DATA_BLOCK "DB_SDC_EMS_HMI"   // DB3814
{ S7_Optimized_Access := 'FALSE' }
VERSION : 0.1
   VAR
      HEADER : Struct
         DB_NR : Int := 3814;
         Res020 : Int := 0;
         Res040 : Int := 0;
         START_EMS : Int := 20;
         LAENGE_EMS : Int := 260;
         OFFSET_EMS_SEK_STAT : Int := 164;
         LAENGE_EMS_SEK_STAT : Int := 34;
         OFFSET_EMS_FKT : Int := 216;
         START_HMI : Int := 20;
         OFFEST_HMI_DATA : Int := 20;
      END_STRUCT;
      HMI : Array[1..30] of Struct
         PULT_Nr_EDIT : Int;
         BILD_Nr : Int;
         BILD_Nr_Alt : Int;
         EMS_Nr : Int;
         EMS_Nr_Alt : Int;
         PROFIL_Nr : Int;
         PROFIL_Nr_Alt : Int;
         Res140 : Int;
         Res160 : Int;
         T_EDIT : Bool;
         T_RESET_BED : Bool;
         T_SAVE : Bool;
         T_LOAD : Bool;
         Res084 : Bool;
         Res085 : Bool;
         Res086 : Bool;
         Res087 : Bool;
         FR_EDIT : Bool;
         ER_DATA : Bool;
         EMS : "UDT_SDC_EMS";
      END_STRUCT;
   END_VAR
BEGIN
   HMI[1].PULT_Nr_EDIT := 0;
   HMI[1].BILD_Nr := 0;
   HMI[1].BILD_Nr_Alt := 0;
   HMI[1].EMS_Nr := 1;
   HMI[1].EMS_Nr_Alt := 1;
   HMI[1].PROFIL_Nr := 0;
   HMI[1].PROFIL_Nr_Alt := 0;
   HMI[1].Res140 := 0;
   HMI[1].Res160 := 0;
   HMI[1].T_EDIT := FALSE;
   HMI[1].T_RESET_BED := FALSE;
   HMI[1].T_SAVE := FALSE;
   HMI[1].T_LOAD := FALSE;
   HMI[1].Res084 := FALSE;
   HMI[1].Res085 := FALSE;
   HMI[1].Res086 := FALSE;
   HMI[1].Res087 := FALSE;
   HMI[1].FR_EDIT := FALSE;
   HMI[1].ER_DATA := FALSE;
   HMI[1].EMS.IF_I_EMS.STAT.LIFE_BIT := FALSE;
   HMI[1].EMS.IF_I_EMS.STAT.ER_SUM := FALSE;
   HMI[1].EMS.IF_I_EMS.STAT.IR_MAN := TRUE;
   HMI[1].EMS.IF_I_EMS.STAT.ER_RESET := FALSE;
   HMI[1].EMS.IF_I_EMS.STAT.HOIST_CLEAR := FALSE;
   HMI[1].EMS.IF_I_EMS.STAT.POS_START_X := FALSE;
   HMI[1].EMS.IF_I_EMS.STAT.ALWAYS_ONE := TRUE;
   HMI[1].EMS.IF_I_EMS.STAT.H_DISABLED := TRUE;
   HMI[1].EMS.IF_I_EMS.STAT.D_FWD := FALSE;
   HMI[1].EMS.IF_I_EMS.STAT.D_RWD := FALSE;
   HMI[1].EMS.IF_I_EMS.STAT.bit12 := FALSE;
   HMI[1].EMS.IF_I_EMS.STAT.D_IN_POS := TRUE;
   HMI[1].EMS.IF_I_EMS.STAT.H_UP := FALSE;
   HMI[1].EMS.IF_I_EMS.STAT.H_DOWN := FALSE;
   HMI[1].EMS.IF_I_EMS.STAT.H_IN_POS := TRUE;
   HMI[1].EMS.IF_I_EMS.STAT.H_IN_TOPPOS := TRUE;
   HMI[1].EMS.IF_I_EMS.STAT.bit2_0 := FALSE;
   HMI[1].EMS.IF_I_EMS.STAT.bit2_1 := FALSE;
   HMI[1].EMS.IF_I_EMS.STAT.bit2_2 := FALSE;
   HMI[1].EMS.IF_I_EMS.STAT.bit2_3 := TRUE;
   HMI[1].EMS.IF_I_EMS.STAT.IN_BOTPOS := FALSE;
   HMI[1].EMS.IF_I_EMS.STAT.bit2_5 := FALSE;
   HMI[1].EMS.IF_I_EMS.STAT.bit2_6 := FALSE;
   HMI[1].EMS.IF_I_EMS.STAT.bit2_7 := FALSE;
   HMI[1].EMS.IF_I_EMS.STAT.MESS_ACT := TRUE;
   HMI[1].EMS.IF_I_EMS.STAT.MESS_POS := FALSE;
   HMI[1].EMS.IF_I_EMS.STAT.bit3_2 := FALSE;
   HMI[1].EMS.IF_I_EMS.STAT.bit3_3 := FALSE;
   HMI[1].EMS.IF_I_EMS.STAT.bit3_4 := FALSE;
   HMI[1].EMS.IF_I_EMS.STAT.bit3_5 := FALSE;
   HMI[1].EMS.IF_I_EMS.STAT.bit3_6 := FALSE;
   HMI[1].EMS.IF_I_EMS.STAT.DATA_TRANS := TRUE;
   HMI[1].EMS.IF_I_EMS.ERROR := 823;
   HMI[1].EMS.IF_I_EMS.D_POS := 466599;
   HMI[1].EMS.IF_I_EMS.H_POS := 4151;
   HMI[1].EMS.IF_I_EMS.VFC.VFC_No := 16#03;
   HMI[1].EMS.IF_I_EMS.VFC.PW1 := 16#EB40;
   HMI[1].EMS.IF_I_EMS.VFC.PW2 := 16#0000;
   HMI[1].EMS.IF_I_EMS.VFC.PW3 := 16#0000;
   HMI[1].EMS.IF_I_EMS.IQ.BS1PH1_KANAL_1 := FALSE;
   HMI[1].EMS.IF_I_EMS.IQ.BS1PH1_KANAL_2 := FALSE;
   HMI[1].EMS.IF_I_EMS.IQ.BS1PH1_KANAL_3 := FALSE;
   HMI[1].EMS.IF_I_EMS.IQ.BS1PH1_KANAL_4 := FALSE;
   HMI[1].EMS.IF_I_EMS.IQ.BS1PH1_KANAL_5 := FALSE;
   HMI[1].EMS.IF_I_EMS.IQ.BS1PH1_KANAL_6 := FALSE;
   HMI[1].EMS.IF_I_EMS.IQ.BS1PH1_KANAL_7 := FALSE;
   HMI[1].EMS.IF_I_EMS.IQ.BS1PH1_KANAL_8 := FALSE;
   HMI[1].EMS.IF_I_EMS.IQ.BS1FC302 := TRUE;
   HMI[1].EMS.IF_I_EMS.IQ.AB1FCM1 := FALSE;
   HMI[1].EMS.IF_I_EMS.IQ.AB1QA1_R := FALSE;
   HMI[1].EMS.IF_I_EMS.IQ.I_1_3 := FALSE;
   HMI[1].EMS.IF_I_EMS.IQ.I_1_8 := FALSE;
   HMI[1].EMS.IF_I_EMS.IQ.I_1_5 := FALSE;
   HMI[1].EMS.IF_I_EMS.IQ.I_1_6 := FALSE;
   HMI[1].EMS.IF_I_EMS.IQ.I_1_7 := FALSE;
   HMI[1].EMS.IF_I_EMS.IQ.HE1BGS03a := TRUE;
   HMI[1].EMS.IF_I_EMS.IQ.HE1BGS03b := TRUE;
   HMI[1].EMS.IF_I_EMS.IQ.HE1BGS05 := TRUE;
   HMI[1].EMS.IF_I_EMS.IQ.BS1SFWE2 := FALSE;
   HMI[1].EMS.IF_I_EMS.IQ.I_2_4 := FALSE;
   HMI[1].EMS.IF_I_EMS.IQ.I_2_5 := FALSE;
   HMI[1].EMS.IF_I_EMS.IQ.I_2_6 := FALSE;
   HMI[1].EMS.IF_I_EMS.IQ.I_2_7 := FALSE;
   HMI[1].EMS.IF_I_EMS.IQ.I_6_0 := FALSE;
   HMI[1].EMS.IF_I_EMS.IQ.I_6_1 := FALSE;
   HMI[1].EMS.IF_I_EMS.IQ.I_6_2 := FALSE;
   HMI[1].EMS.IF_I_EMS.IQ.I_6_3 := FALSE;
   HMI[1].EMS.IF_I_EMS.IQ.I_6_4 := FALSE;
   HMI[1].EMS.IF_I_EMS.IQ.I_6_5 := FALSE;
   HMI[1].EMS.IF_I_EMS.IQ.I_6_6 := FALSE;
   HMI[1].EMS.IF_I_EMS.IQ.I_6_7 := FALSE;
   HMI[1].EMS.IF_I_EMS.IQ."BS1PH1_L+" := TRUE;
   HMI[1].EMS.IF_I_EMS.IQ.BS1PH1_DAT := FALSE;
   HMI[1].EMS.IF_I_EMS.IQ.AB1QA1 := FALSE;
   HMI[1].EMS.IF_I_EMS.IQ.O_0_3 := FALSE;
   HMI[1].EMS.IF_I_EMS.IQ.O_0_4 := FALSE;
   HMI[1].EMS.IF_I_EMS.IQ.O_0_5 := FALSE;
   HMI[1].EMS.IF_I_EMS.IQ.O_0_6 := FALSE;
   HMI[1].EMS.IF_I_EMS.IQ.O_0_7 := FALSE;
   HMI[1].EMS.IF_I_EMS.IQ.HE1KK1 := FALSE;
   HMI[1].EMS.IF_I_EMS.IQ.O_8_1 := FALSE;
   HMI[1].EMS.IF_I_EMS.IQ.O_8_2 := FALSE;
   HMI[1].EMS.IF_I_EMS.IQ.O_8_3 := FALSE;
   HMI[1].EMS.IF_I_EMS.IQ.O_8_4 := FALSE;
   HMI[1].EMS.IF_I_EMS.IQ.O_8_5 := FALSE;
   HMI[1].EMS.IF_I_EMS.IQ.O_8_6 := FALSE;
   HMI[1].EMS.IF_I_EMS.IQ.O_8_7 := FALSE;
   HMI[1].EMS.IF_I_EMS.IQ.I_261_0 := FALSE;
   HMI[1].EMS.IF_I_EMS.IQ.I_261_1 := FALSE;
   HMI[1].EMS.IF_I_EMS.IQ.I_261_2 := FALSE;
   HMI[1].EMS.IF_I_EMS.IQ.I_261_3 := FALSE;
   HMI[1].EMS.IF_I_EMS.IQ.I_261_4 := FALSE;
   HMI[1].EMS.IF_I_EMS.IQ.I_261_5 := FALSE;
   HMI[1].EMS.IF_I_EMS.IQ.I_261_6 := FALSE;
   HMI[1].EMS.IF_I_EMS.IQ.I_261_7 := FALSE;
   HMI[1].EMS.IF_I_EMS.IQ.HE1BGG1 := TRUE;
   HMI[1].EMS.IF_I_EMS.IQ."HE1BGG1:13" := FALSE;
   HMI[1].EMS.IF_I_EMS.IQ.HE1BGE05 := TRUE;
   HMI[1].EMS.IF_I_EMS.IQ.I_271_3 := FALSE;
   HMI[1].EMS.IF_I_EMS.IQ.I_271_4 := FALSE;
   HMI[1].EMS.IF_I_EMS.IQ.I_271_5 := FALSE;
   HMI[1].EMS.IF_I_EMS.IQ.I_271_6 := FALSE;
   HMI[1].EMS.IF_I_EMS.IQ.I_271_7 := FALSE;
   HMI[1].EMS.IF_I_EMS.IQ.SN1BGE04 := TRUE;
   HMI[1].EMS.IF_I_EMS.IQ.I_281_1 := FALSE;
   HMI[1].EMS.IF_I_EMS.IQ.I_281_2 := FALSE;
   HMI[1].EMS.IF_I_EMS.IQ.I_281_3 := FALSE;
   HMI[1].EMS.IF_I_EMS.IQ.I_281_4 := FALSE;
   HMI[1].EMS.IF_I_EMS.IQ.I_281_5 := FALSE;
   HMI[1].EMS.IF_I_EMS.IQ.I_281_6 := FALSE;
   HMI[1].EMS.IF_I_EMS.IQ.I_281_7 := FALSE;
   HMI[1].EMS.IF_I_EMS.IQ.I_285_0 := FALSE;
   HMI[1].EMS.IF_I_EMS.IQ.I_285_1 := FALSE;
   HMI[1].EMS.IF_I_EMS.IQ.I_285_2 := FALSE;
   HMI[1].EMS.IF_I_EMS.IQ.I_285_3 := FALSE;
   HMI[1].EMS.IF_I_EMS.IQ.I_285_4 := FALSE;
   HMI[1].EMS.IF_I_EMS.IQ.I_285_5 := FALSE;
   HMI[1].EMS.IF_I_EMS.IQ.I_285_6 := FALSE;
   HMI[1].EMS.IF_I_EMS.IQ.I_285_7 := FALSE;
   HMI[1].EMS.IF_I_EMS.ER_WORD_No := 25;
   HMI[1].EMS.IF_I_EMS.ER_WORD := 16#0002;
   HMI[1].EMS.IF_I_EMS.FB_DBNo := 2;
   HMI[1].EMS.IF_I_EMS.FB_DBBNo := 20;
   HMI[1].EMS.IF_Q_EMS.EMS_ID := 1;
   HMI[1].EMS.IF_Q_EMS.CONT.LIFE_BIT := TRUE;
   HMI[1].EMS.IF_Q_EMS.CONT.ER_SDC := FALSE;
   HMI[1].EMS.IF_Q_EMS.CONT.H_EMERG := FALSE;
   HMI[1].EMS.IF_Q_EMS.CONT.Spare_0_3 := FALSE;
   HMI[1].EMS.IF_Q_EMS.CONT.LAMP_TEST := FALSE;
   HMI[1].EMS.IF_Q_EMS.CONT.VAC_CLEAN := FALSE;
   HMI[1].EMS.IF_Q_EMS.CONT.SYNCH := FALSE;
   HMI[1].EMS.IF_Q_EMS.CONT.DATA_TRANS := TRUE;
   HMI[1].EMS.IF_Q_EMS.CONT.ER_RESET := FALSE;
   HMI[1].EMS.IF_Q_EMS.CONT.AUTO := FALSE;
   HMI[1].EMS.IF_Q_EMS.CONT.MAN := TRUE;
   HMI[1].EMS.IF_Q_EMS.CONT.D_C_BREAK := FALSE;
   HMI[1].EMS.IF_Q_EMS.CONT.H_C_BREAK := FALSE;
   HMI[1].EMS.IF_Q_EMS.CONT.D_EMERG_FC := FALSE;
   HMI[1].EMS.IF_Q_EMS.CONT.INC_TOL_POS := FALSE;
   HMI[1].EMS.IF_Q_EMS.CONT.E_STOP := FALSE;
   HMI[1].EMS.IF_Q_EMS.CONT.D_C_FWD := FALSE;
   HMI[1].EMS.IF_Q_EMS.CONT.D_C_RWD := FALSE;
   HMI[1].EMS.IF_Q_EMS.CONT.D_C_BSP := FALSE;
   HMI[1].EMS.IF_Q_EMS.CONT.Spare_2_3 := FALSE;
   HMI[1].EMS.IF_Q_EMS.CONT.IR_noEMSnumber := FALSE;
   HMI[1].EMS.IF_Q_EMS.CONT.IR_noLogin := FALSE;
   HMI[1].EMS.IF_Q_EMS.CONT.BYP_scalance_PN_error := FALSE;
   HMI[1].EMS.IF_Q_EMS.CONT.Spare_2_7 := FALSE;
   HMI[1].EMS.IF_Q_EMS.CONT.H_C_UP := FALSE;
   HMI[1].EMS.IF_Q_EMS.CONT.H_C_DOWN := FALSE;
   HMI[1].EMS.IF_Q_EMS.CONT.H_C_POS := FALSE;
   HMI[1].EMS.IF_Q_EMS.CONT.H_C_TOP := FALSE;
   HMI[1].EMS.IF_Q_EMS.CONT.H_EN := TRUE;
   HMI[1].EMS.IF_Q_EMS.CONT.H_BYP_ROPE := FALSE;
   HMI[1].EMS.IF_Q_EMS.CONT.Spare_3_6 := FALSE;
   HMI[1].EMS.IF_Q_EMS.CONT.H_BYP_REF_INI := FALSE;
   HMI[1].EMS.IF_Q_EMS.D_SETPOS := 466601;
   HMI[1].EMS.IF_Q_EMS.D_SETSPEED := 4000;
   HMI[1].EMS.IF_Q_EMS.H_SETPOS := 4151;
   HMI[1].EMS.IF_Q_EMS.H_SETSPEED := 0;
   HMI[1].EMS.IF_Q_EMS.FB_VFC_No := 16#03;
   HMI[1].EMS.IF_Q_EMS.FB_ER_WORD_No := 25;
   HMI[1].EMS.IF_Q_EMS.DB_No := 2;
   HMI[1].EMS.IF_Q_EMS.DBB_No := 24;
   HMI[1].EMS.IF_Q_EMS.DB_UserData := 16#2710_3B1A;
   HMI[1].EMS.IF_Q_EMS.ERRORS_SPLC._901_ER_SUM := FALSE;
   HMI[1].EMS.IF_Q_EMS.ERRORS_SPLC._902_ER_SUM_SDC := FALSE;
   HMI[1].EMS.IF_Q_EMS.ERRORS_SPLC._903_ER_BC_JUMP := FALSE;
   HMI[1].EMS.IF_Q_EMS.ERRORS_SPLC._904_ER_NO_SEK := FALSE;
   HMI[1].EMS.IF_Q_EMS.ERRORS_SPLC._905_ER_COMMAND := FALSE;
   HMI[1].EMS.IF_Q_EMS.ERRORS_SPLC._906_ER_BC_LIM := FALSE;
   HMI[1].EMS.IF_Q_EMS.ERRORS_SPLC._907_ER_EMS_ID := FALSE;
   HMI[1].EMS.IF_Q_EMS.ERRORS_SPLC._908_ER_SEK_NR := FALSE;
   HMI[1].EMS.IF_Q_EMS.ERRORS_SPLC._909_ER_LIFE := FALSE;
   HMI[1].EMS.IF_Q_EMS.ERRORS_SPLC._910_ER_BUS := FALSE;
   HMI[1].EMS.IF_Q_EMS.ERRORS_SPLC._911 := FALSE;
   HMI[1].EMS.IF_Q_EMS.ERRORS_SPLC._912 := FALSE;
   HMI[1].EMS.IF_Q_EMS.ERRORS_SPLC._913 := FALSE;
   HMI[1].EMS.IF_Q_EMS.ERRORS_SPLC._914 := FALSE;
   HMI[1].EMS.IF_Q_EMS.ERRORS_SPLC._915 := FALSE;
   HMI[1].EMS.IF_Q_EMS.ERRORS_SPLC._916 := FALSE;
   // 9920 more start values not shown
END_DATA_BLOCK

DATA_BLOCK "DB_SDC_TS_IF_HMI"   // DB3816
{ S7_Optimized_Access := 'FALSE' }
AUTHOR : FFM
FAMILY : SDC
NAME : SECT_DEF
VERSION : 1.0
   VAR
      HEADER : Struct
         DB_NR : Int := 3816;
         Res020 : Int := 0;
         Res040 : Int := 0;
         START_DAT : Int := 1;
         LAENGE_SEK_COM : Int := 18;
         LAENGE_SEK_STAT : Int := 34;
         OFFEST_SEK_STAT : Int := 18;
         Res140 : Int := 44;
         START_HMI : Int := 20;
         OFFEST_HMI_DATA : Int := 20;
      END_STRUCT;
      HMI : Array[1..30] of Struct
         PULT_Nr_EDIT : Int;
         BILD_Nr : Int;
         BILD_Nr_Alt : Int;
         SEK_Nr : Int;
         SEK_Nr_Alt : Int;
         Res100 : Int;
         Res120 : Int;
         Res140 : Int;
         Res160 : Int;
         T_EDIT : Bool;
         T_RESET_BED : Bool;
         T_SAVE : Bool;
         T_LOAD : Bool;
         Res084 : Bool;
         Res085 : Bool;
         Res086 : Bool;
         Res087 : Bool;
         FR_EDIT : Bool;
         ER_DATA : Bool;
         COM : "UDT_SDC_EMS_TS_COM";
         STAT : "UDT_SDC_EMS_TS_STAT";
      END_STRUCT;
   END_VAR
BEGIN
   HMI[1].PULT_Nr_EDIT := 0;
   HMI[1].BILD_Nr := 0;
   HMI[1].BILD_Nr_Alt := 0;
   HMI[1].SEK_Nr := 1;
   HMI[1].SEK_Nr_Alt := 255;
   HMI[1].Res100 := 0;
   HMI[1].Res120 := 0;
   HMI[1].Res140 := 0;
   HMI[1].Res160 := 0;
   HMI[1].T_EDIT := FALSE;
   HMI[1].T_RESET_BED := FALSE;
   HMI[1].T_SAVE := FALSE;
   HMI[1].T_LOAD := FALSE;
   HMI[1].Res084 := FALSE;
   HMI[1].Res085 := FALSE;
   HMI[1].Res086 := FALSE;
   HMI[1].Res087 := FALSE;
   HMI[1].FR_EDIT := FALSE;
   HMI[1].ER_DATA := FALSE;
   HMI[1].COM.VAL.PROFIL := 0;
   HMI[1].COM.VAL.D_SETSPEED := 0;
   HMI[1].COM.VAL.D_POS_OFFS := 0;
   HMI[1].COM.BIT.ER_RESET := FALSE;
   HMI[1].COM.BIT.AUTO := FALSE;
   HMI[1].COM.BIT.MAN := FALSE;
   HMI[1].COM.BIT.Spare_0_3 := FALSE;
   HMI[1].COM.BIT.Spare_0_4 := FALSE;
   HMI[1].COM.BIT.E_STOP := TRUE;
   HMI[1].COM.BIT.Spare_0_6 := FALSE;
   HMI[1].COM.BIT.Spare_0_7 := FALSE;
   HMI[1].COM.BIT.D_C_FWD := FALSE;
   HMI[1].COM.BIT.D_C_RWD := FALSE;
   HMI[1].COM.BIT.D_C_BSP := FALSE;
   HMI[1].COM.BIT.D_C_V1 := TRUE;
   HMI[1].COM.BIT.D_C_V2 := FALSE;
   HMI[1].COM.BIT.D_C_V_VAR := FALSE;
   HMI[1].COM.BIT.D_C_BEFOR_POS := FALSE;
   HMI[1].COM.BIT.D_C_AFTER_POS := FALSE;
   HMI[1].COM.BIT.H_C_RAISE := FALSE;
   HMI[1].COM.BIT.H_C_LOWER := FALSE;
   HMI[1].COM.BIT.H_C_POS := FALSE;
   HMI[1].COM.BIT.H_C_POS1 := FALSE;
   HMI[1].COM.BIT.H_C_POS2 := FALSE;
   HMI[1].COM.BIT.H_C_POS3 := FALSE;
   HMI[1].COM.BIT.H_C_POS4 := FALSE;
   HMI[1].COM.BIT.H_C_TOP := FALSE;
   HMI[1].COM.BIT.H_BYP_ROPE := FALSE;
   HMI[1].COM.BIT.Spare_3_1 := FALSE;
   HMI[1].COM.BIT.H_BYP_REF_INI := FALSE;
   HMI[1].COM.BIT.H_C_SLOW := FALSE;
   HMI[1].COM.BIT.D_BYP_DIST_CONTR := FALSE;
   HMI[1].COM.BIT.Spare_3_5 := FALSE;
   HMI[1].COM.BIT.Spare_3_6 := FALSE;
   HMI[1].COM.BIT.SET_PROF := FALSE;
   HMI[1].COM.FKT_SET.EMS_TO_REPAIR_1 := FALSE;
   HMI[1].COM.FKT_SET.EMS_TO_REPAIR_2 := FALSE;
   HMI[1].COM.FKT_SET.EMERG_HOIST := FALSE;
   HMI[1].COM.FKT_SET.Reserve_03 := FALSE;
   HMI[1].COM.FKT_SET.EMERG_DRIVE_FC := FALSE;
   HMI[1].COM.FKT_SET.Reserve_05 := FALSE;
   HMI[1].COM.FKT_SET.LAMP_TEST := FALSE;
   HMI[1].COM.FKT_SET.VAC_CLEAN := FALSE;
   HMI[1].COM.FKT_SET.PE_TEST := FALSE;
   HMI[1].COM.FKT_SET.KOHLE_TEST := FALSE;
   HMI[1].COM.FKT_SET.KOM_TEST := FALSE;
   HMI[1].COM.FKT_SET.Reserve_11 := FALSE;
   HMI[1].COM.FKT_SET.Reserve_12 := FALSE;
   HMI[1].COM.FKT_SET.Reserve_13 := FALSE;
   HMI[1].COM.FKT_SET.Reserve_14 := FALSE;
   HMI[1].COM.FKT_SET.Reserve_15 := FALSE;
   HMI[1].COM.FKT_RESET.EMS_TO_REPAIR_1 := FALSE;
   HMI[1].COM.FKT_RESET.EMS_TO_REPAIR_2 := FALSE;
   HMI[1].COM.FKT_RESET.EMERG_HOIST := FALSE;
   HMI[1].COM.FKT_RESET.Reserve_03 := FALSE;
   HMI[1].COM.FKT_RESET.EMERG_DRIVE_FC := FALSE;
   HMI[1].COM.FKT_RESET.Reserve_05 := FALSE;
   HMI[1].COM.FKT_RESET.LAMP_TEST := FALSE;
   HMI[1].COM.FKT_RESET.VAC_CLEAN := FALSE;
   HMI[1].COM.FKT_RESET.PE_TEST := FALSE;
   HMI[1].COM.FKT_RESET.KOHLE_TEST := FALSE;
   HMI[1].COM.FKT_RESET.KOM_TEST := FALSE;
   HMI[1].COM.FKT_RESET.Reserve_11 := FALSE;
   HMI[1].COM.FKT_RESET.Reserve_12 := FALSE;
   HMI[1].COM.FKT_RESET.Reserve_13 := FALSE;
   HMI[1].COM.FKT_RESET.Reserve_14 := FALSE;
   HMI[1].COM.FKT_RESET.Reserve_15 := FALSE;
   HMI[1].STAT.VAL.EMS_ID := 9;
   HMI[1].STAT.VAL.PROFIL := 1;
   HMI[1].STAT.VAL.DRIVE_POS := 27823;
   HMI[1].STAT.VAL.HOIST_POS := 2747;
   HMI[1].STAT.VAL.ERROR := 824;
   HMI[1].STAT.VAL.DRIVE_POS_PERC := 51;
   HMI[1].STAT.VAL.SEK := 255;
   HMI[1].STAT.BIT.PRESENT := TRUE;
   HMI[1].STAT.BIT.ERROR := FALSE;
   HMI[1].STAT.BIT.MAN_IR := FALSE;
   HMI[1].STAT.BIT.MORE_EMS_PRESENT := FALSE;
   HMI[1].STAT.BIT.ER_COMMAND := FALSE;
   HMI[1].STAT.BIT.W_DIST := FALSE;
   HMI[1].STAT.BIT.Spare_0_6 := FALSE;
   HMI[1].STAT.BIT.MESS_ACT := TRUE;
   HMI[1].STAT.BIT.D_MOVING := FALSE;
   HMI[1].STAT.BIT.D_NOT_MOVING := TRUE;
   HMI[1].STAT.BIT.H_MOVING := FALSE;
   HMI[1].STAT.BIT.H_NOT_MOVING := TRUE;
   HMI[1].STAT.BIT.X_MOVING := FALSE;
   HMI[1].STAT.BIT.X_NOT_MOVING := TRUE;
   HMI[1].STAT.BIT.D_IN_POS := TRUE;
   HMI[1].STAT.BIT.Spare_2_1 := FALSE;
   HMI[1].STAT.BIT.D_BEFOR_POS := FALSE;
   HMI[1].STAT.BIT.D_AFTER_POS := FALSE;
   HMI[1].STAT.BIT.D_GR_AP1 := TRUE;
   HMI[1].STAT.BIT.D_SM_AP1 := FALSE;
   HMI[1].STAT.BIT.D_GR_AP2 := TRUE;
   HMI[1].STAT.BIT.D_SM_AP2 := FALSE;
   HMI[1].STAT.BIT.H_IN_POS := TRUE;
   HMI[1].STAT.BIT.H_IN_TOPPOS := FALSE;
   HMI[1].STAT.BIT.H_IN_POS1 := TRUE;
   HMI[1].STAT.BIT.H_IN_POS2 := TRUE;
   HMI[1].STAT.BIT.H_IN_POS3 := TRUE;
   HMI[1].STAT.BIT.H_IN_POS4 := TRUE;
   HMI[1].STAT.BIT.H_GR_POS := FALSE;
   HMI[1].STAT.BIT.H_SM_POS := FALSE;
   HMI[1].STAT.BIT.H_GR_POS1 := FALSE;
   HMI[1].STAT.BIT.H_SM_POS1 := FALSE;
   HMI[1].STAT.BIT.H_GR_POS2 := FALSE;
   HMI[1].STAT.BIT.H_SM_POS2 := FALSE;
   HMI[1].STAT.BIT.H_GR_POS3 := FALSE;
   HMI[1].STAT.BIT.H_SM_POS3 := FALSE;
   HMI[1].STAT.BIT.H_GR_POS4 := FALSE;
   HMI[1].STAT.BIT.H_SM_POS4 := FALSE;
   HMI[1].STAT.BIT.H_BOTTOM_POS := FALSE;
   HMI[1].STAT.BIT.H_DISABLED := FALSE;
   HMI[1].STAT.BIT.H_CLEAR := FALSE;
   HMI[1].STAT.BIT.D_MOVING_FWD := FALSE;
   HMI[1].STAT.BIT.D_MOVING_RWD := FALSE;
   HMI[1].STAT.BIT.D_RESET_AFTER := FALSE;
   HMI[1].STAT.BIT.D_PULK := FALSE;
   HMI[1].STAT.BIT.D_NO_POS := FALSE;
   HMI[1].STAT.SORTE[1] := 'L';
   HMI[1].STAT.SORTE[2] := 'E';
   HMI[1].STAT.SORTE[3] := 'E';
   HMI[1].STAT.SORTE[4] := 'R';
   HMI[1].STAT.FKT.EMS_TO_REPAIR_1 := FALSE;
   HMI[1].STAT.FKT.EMS_TO_REPAIR_2 := FALSE;
   HMI[1].STAT.FKT.EMERG_HOIST := FALSE;
   HMI[1].STAT.FKT.Reserve_03 := FALSE;
   HMI[1].STAT.FKT.EMERG_DRIVE_FC := FALSE;
   HMI[1].STAT.FKT.Reserve_05 := FALSE;
   HMI[1].STAT.FKT.LAMP_TEST := FALSE;
   HMI[1].STAT.FKT.VAC_CLEAN := FALSE;
   HMI[1].STAT.FKT.PE_TEST := FALSE;
   HMI[1].STAT.FKT.KOHLE_TEST := FALSE;
   HMI[1].STAT.FKT.KOM_TEST := FALSE;
   HMI[1].STAT.FKT.Reserve_11 := FALSE;
   HMI[1].STAT.FKT.Reserve_12 := FALSE;
   HMI[1].STAT.FKT.Reserve_13 := FALSE;
   HMI[1].STAT.FKT.Reserve_14 := FALSE;
   HMI[1].STAT.FKT.Reserve_15 := FALSE;
   HMI[1].STAT.SPARE := 16#0000;
   HMI[2].PULT_Nr_EDIT := 0;
   HMI[2].BILD_Nr := 0;
   HMI[2].BILD_Nr_Alt := 0;
   HMI[2].SEK_Nr := 1;
   HMI[2].SEK_Nr_Alt := 262;
   HMI[2].Res100 := 0;
   HMI[2].Res120 := 0;
   HMI[2].Res140 := 0;
   HMI[2].Res160 := 0;
   HMI[2].T_EDIT := FALSE;
   HMI[2].T_RESET_BED := FALSE;
   HMI[2].T_SAVE := FALSE;
   HMI[2].T_LOAD := FALSE;
   HMI[2].Res084 := FALSE;
   HMI[2].Res085 := FALSE;
   HMI[2].Res086 := FALSE;
   HMI[2].Res087 := FALSE;
   HMI[2].FR_EDIT := FALSE;
   HMI[2].ER_DATA := FALSE;
   HMI[2].COM.VAL.PROFIL := 0;
   HMI[2].COM.VAL.D_SETSPEED := 0;
   HMI[2].COM.VAL.D_POS_OFFS := 0;
   HMI[2].COM.BIT.ER_RESET := FALSE;
   HMI[2].COM.BIT.AUTO := TRUE;
   HMI[2].COM.BIT.MAN := FALSE;
   HMI[2].COM.BIT.Spare_0_3 := FALSE;
   HMI[2].COM.BIT.Spare_0_4 := FALSE;
   HMI[2].COM.BIT.E_STOP := FALSE;
   HMI[2].COM.BIT.Spare_0_6 := FALSE;
   HMI[2].COM.BIT.Spare_0_7 := FALSE;
   HMI[2].COM.BIT.D_C_FWD := TRUE;
   HMI[2].COM.BIT.D_C_RWD := FALSE;
   HMI[2].COM.BIT.D_C_BSP := TRUE;
   HMI[2].COM.BIT.D_C_V1 := TRUE;
   HMI[2].COM.BIT.D_C_V2 := FALSE;
   HMI[2].COM.BIT.D_C_V_VAR := FALSE;
   HMI[2].COM.BIT.D_C_BEFOR_POS := TRUE;
   HMI[2].COM.BIT.D_C_AFTER_POS := TRUE;
   HMI[2].COM.BIT.H_C_RAISE := FALSE;
   HMI[2].COM.BIT.H_C_LOWER := FALSE;
   // 3000 more start values not shown
END_DATA_BLOCK

// folder: 06_IDBs

DATA_BLOCK "IDB504_ZONE_5"   // DB13
{ S7_Optimized_Access := 'FALSE' }
VERSION : 0.1
"FB115_FB_Zone"
BEGIN
END_DATA_BLOCK

DATA_BLOCK "IDB501_ZONE_1"   // DB501
{ S7_Optimized_Access := 'FALSE' }
VERSION : 0.1
"FB115_FB_Zone"
BEGIN
END_DATA_BLOCK

DATA_BLOCK "IDB502_ZONE_2"   // DB502
{ S7_Optimized_Access := 'FALSE' }
VERSION : 0.1
"FB115_FB_Zone"
BEGIN
END_DATA_BLOCK

DATA_BLOCK "IDB503_ZONE_3"   // DB503
{ S7_Optimized_Access := 'FALSE' }
VERSION : 0.1
"FB115_FB_Zone"
BEGIN
END_DATA_BLOCK

DATA_BLOCK "IDB504_ZONE_4"   // DB504
{ S7_Optimized_Access := 'FALSE' }
VERSION : 0.1
"FB115_FB_Zone"
BEGIN
END_DATA_BLOCK

DATA_BLOCK "IDB505_ZONE_5"   // DB505
{ S7_Optimized_Access := 'FALSE' }
VERSION : 0.1
"FB115_FB_Zone"
BEGIN
END_DATA_BLOCK

DATA_BLOCK "IDB506_ZONE_6"   // DB506
{ S7_Optimized_Access := 'FALSE' }
VERSION : 0.1
"FB115_FB_Zone"
BEGIN
END_DATA_BLOCK

DATA_BLOCK "IDB543_ZONE_43"   // DB543
{ S7_Optimized_Access := 'FALSE' }
VERSION : 0.1
"FB115_FB_Zone"
BEGIN
END_DATA_BLOCK

DATA_BLOCK "IDB544_ZONE_44"   // DB544
{ S7_Optimized_Access := 'FALSE' }
VERSION : 0.1
"FB115_FB_Zone"
BEGIN
END_DATA_BLOCK

DATA_BLOCK "IDB547_ZONE_47"   // DB547
{ S7_Optimized_Access := 'FALSE' }
VERSION : 0.1
"FB115_FB_Zone"
BEGIN
END_DATA_BLOCK

DATA_BLOCK "IDB548_ZONE_48"   // DB548
{ S7_Optimized_Access := 'FALSE' }
VERSION : 0.1
"FB115_FB_Zone"
BEGIN
END_DATA_BLOCK

DATA_BLOCK "IDB552_ZONE_52"   // DB552
{ S7_Optimized_Access := 'FALSE' }
VERSION : 0.1
"FB115_FB_Zone"
BEGIN
END_DATA_BLOCK

DATA_BLOCK "IDB558_ZONE_58"   // DB558
{ S7_Optimized_Access := 'FALSE' }
VERSION : 0.1
"FB115_FB_Zone"
BEGIN
END_DATA_BLOCK

DATA_BLOCK "IDB600_ZonePositionArrayTrafficCop_DB"   // DB600
{ S7_Optimized_Access := 'FALSE' }
VERSION : 0.1
"FB116_FB_ZonePositionArrayTrafficCop"
BEGIN
END_DATA_BLOCK

DATA_BLOCK "IDB601_MapSDCOut_Carrier_DB"   // DB601
{ S7_Optimized_Access := 'TRUE' }
VERSION : 0.1
"FB117_MapSDCOut_Carrier"
BEGIN
END_DATA_BLOCK

DATA_BLOCK "IDB602_NextCarrierTCopMotionFB"   // DB602
{ S7_Optimized_Access := 'TRUE' }
VERSION : 0.1
"FB111_NextCarrierTCopMotionFB"
BEGIN
END_DATA_BLOCK

DATA_BLOCK "IDB603_FB_ZonePositionArrayTrafficCop_DB"   // DB603
{ S7_Optimized_Access := 'FALSE' }
VERSION : 0.1
"FB116_FB_ZonePositionArrayTrafficCop"
BEGIN
END_DATA_BLOCK

DATA_BLOCK "IDB604_SpacingCheck"   // DB604
{ S7_Optimized_Access := 'TRUE' }
VERSION : 0.1
"FB120_ZoneSpacingCheck"
BEGIN
END_DATA_BLOCK

DATA_BLOCK "IDB605_CARRIER"   // DB605
{ S7_Optimized_Access := 'TRUE' }
VERSION : 0.1
"FB112_Carrier"
BEGIN
END_DATA_BLOCK

DATA_BLOCK "IDB606_FirstCarrierTCopMotionFB"   // DB606
{ S7_Optimized_Access := 'TRUE' }
VERSION : 0.1
"FB110_FirstCarrierTCopMotionFB"
BEGIN
END_DATA_BLOCK

DATA_BLOCK "IDB607_FirstCarrierTCopMotionFB"   // DB607
{ S7_Optimized_Access := 'TRUE' }
VERSION : 0.1
"FB110_FirstCarrierTCopMotionFB"
BEGIN
END_DATA_BLOCK

DATA_BLOCK "IDB608_NextCarrierTCopMotionFB"   // DB608
{ S7_Optimized_Access := 'TRUE' }
VERSION : 0.1
"FB111_NextCarrierTCopMotionFB"
BEGIN
END_DATA_BLOCK

DATA_BLOCK "IDB609_TCMapSDCOutFB"   // DB609
{ S7_Optimized_Access := 'TRUE' }
VERSION : 0.1
"FB118_TCMapSDCOut"
BEGIN
END_DATA_BLOCK

DATA_BLOCK "IDB610_SpacingCheckFB"   // DB610
{ S7_Optimized_Access := 'TRUE' }
VERSION : 0.1
"FB120_ZoneSpacingCheck"
BEGIN
END_DATA_BLOCK

// folder: System blocks/Program resources

DATA_BLOCK "Reset_Timer"   // DB1
{ S7_Optimized_Access := 'TRUE' }
AUTHOR : Simatic
FAMILY : IEC
NAME : IEC_TMR
VERSION : 1.0
"IEC_TIMER"
BEGIN
END_DATA_BLOCK

DATA_BLOCK "C23_Heartbeat_On_Timer"   // DB2
{ S7_Optimized_Access := 'TRUE' }
AUTHOR : Simatic
FAMILY : IEC
NAME : IEC_TMR
VERSION : 1.0
"IEC_TIMER"
BEGIN
END_DATA_BLOCK

DATA_BLOCK "EMS_Heartbeat_On_Timer"   // DB3
{ S7_Optimized_Access := 'TRUE' }
AUTHOR : Simatic
FAMILY : IEC
NAME : IEC_TMR
VERSION : 1.0
"IEC_TIMER"
BEGIN
END_DATA_BLOCK

DATA_BLOCK "C23_Heartbeat_Off_Timer"   // DB5
{ S7_Optimized_Access := 'TRUE' }
AUTHOR : Simatic
FAMILY : IEC
NAME : IEC_TMR
VERSION : 1.0
"IEC_TIMER"
BEGIN
END_DATA_BLOCK

DATA_BLOCK "C22_Heartbeat_On_Timer"   // DB6
{ S7_Optimized_Access := 'TRUE' }
AUTHOR : Simatic
FAMILY : IEC
NAME : IEC_TMR
VERSION : 1.0
"IEC_TIMER"
BEGIN
END_DATA_BLOCK

DATA_BLOCK "EMS_Heartbeat_Off_Timer"   // DB7
{ S7_Optimized_Access := 'TRUE' }
AUTHOR : Simatic
FAMILY : IEC
NAME : IEC_TMR
VERSION : 1.0
"IEC_TIMER"
BEGIN
END_DATA_BLOCK

DATA_BLOCK "C22_Heartbeat_Off_Timer"   // DB9
{ S7_Optimized_Access := 'TRUE' }
AUTHOR : Simatic
FAMILY : IEC
NAME : IEC_TMR
VERSION : 1.0
"IEC_TIMER"
BEGIN
END_DATA_BLOCK

DATA_BLOCK "C21_Heartbeat_On_Timer"   // DB10
{ S7_Optimized_Access := 'TRUE' }
AUTHOR : Simatic
FAMILY : IEC
NAME : IEC_TMR
VERSION : 1.0
"IEC_TIMER"
BEGIN
END_DATA_BLOCK

DATA_BLOCK "C21_Heartbeat_Off_Timer"   // DB12
{ S7_Optimized_Access := 'TRUE' }
AUTHOR : Simatic
FAMILY : IEC
NAME : IEC_TMR
VERSION : 1.0
"IEC_TIMER"
BEGIN
END_DATA_BLOCK

DATA_BLOCK "C24_Heartbeat_On_Timer"   // DB17
{ S7_Optimized_Access := 'TRUE' }
AUTHOR : Simatic
FAMILY : IEC
NAME : IEC_TMR
VERSION : 1.0
"IEC_TIMER"
BEGIN
END_DATA_BLOCK

DATA_BLOCK "C24_Heartbeat_Off_Timer"   // DB18
{ S7_Optimized_Access := 'TRUE' }
AUTHOR : Simatic
FAMILY : IEC
NAME : IEC_TMR
VERSION : 1.0
"IEC_TIMER"
BEGIN
END_DATA_BLOCK

DATA_BLOCK "C25_Heartbeat_On_Timer"   // DB19
{ S7_Optimized_Access := 'TRUE' }
AUTHOR : Simatic
FAMILY : IEC
NAME : IEC_TMR
VERSION : 1.0
"IEC_TIMER"
BEGIN
END_DATA_BLOCK

DATA_BLOCK "C25_Heartbeat_Off_Timer"   // DB20
{ S7_Optimized_Access := 'TRUE' }
AUTHOR : Simatic
FAMILY : IEC
NAME : IEC_TMR
VERSION : 1.0
"IEC_TIMER"
BEGIN
END_DATA_BLOCK

DATA_BLOCK "C26_Heartbeat_On_Timer"   // DB21
{ S7_Optimized_Access := 'TRUE' }
AUTHOR : Simatic
FAMILY : IEC
NAME : IEC_TMR
VERSION : 1.0
"IEC_TIMER"
BEGIN
END_DATA_BLOCK

DATA_BLOCK "C26_Heartbeat_Off_Timer"   // DB22
{ S7_Optimized_Access := 'TRUE' }
AUTHOR : Simatic
FAMILY : IEC
NAME : IEC_TMR
VERSION : 1.0
"IEC_TIMER"
BEGIN
END_DATA_BLOCK

DATA_BLOCK "C27_Heartbeat_On_Timer"   // DB23
{ S7_Optimized_Access := 'TRUE' }
AUTHOR : Simatic
FAMILY : IEC
NAME : IEC_TMR
VERSION : 1.0
"IEC_TIMER"
BEGIN
END_DATA_BLOCK

DATA_BLOCK "C27_Heartbeat_Off_Timer"   // DB24
{ S7_Optimized_Access := 'TRUE' }
AUTHOR : Simatic
FAMILY : IEC
NAME : IEC_TMR
VERSION : 1.0
"IEC_TIMER"
BEGIN
END_DATA_BLOCK

DATA_BLOCK "C28_Heartbeat_On_Timer"   // DB25
{ S7_Optimized_Access := 'TRUE' }
AUTHOR : Simatic
FAMILY : IEC
NAME : IEC_TMR
VERSION : 1.0
"IEC_TIMER"
BEGIN
END_DATA_BLOCK

DATA_BLOCK "C28_Heartbeat_Off_Timer"   // DB26
{ S7_Optimized_Access := 'TRUE' }
AUTHOR : Simatic
FAMILY : IEC
NAME : IEC_TMR
VERSION : 1.0
"IEC_TIMER"
BEGIN
END_DATA_BLOCK

DATA_BLOCK "C29_Heartbeat_On_Timer"   // DB27
{ S7_Optimized_Access := 'TRUE' }
AUTHOR : Simatic
FAMILY : IEC
NAME : IEC_TMR
VERSION : 1.0
"IEC_TIMER"
BEGIN
END_DATA_BLOCK

DATA_BLOCK "C29_Heartbeat_Off_Timer"   // DB28
{ S7_Optimized_Access := 'TRUE' }
AUTHOR : Simatic
FAMILY : IEC
NAME : IEC_TMR
VERSION : 1.0
"IEC_TIMER"
BEGIN
END_DATA_BLOCK

DATA_BLOCK "C30_Heartbeat_On_Timer"   // DB29
{ S7_Optimized_Access := 'TRUE' }
AUTHOR : Simatic
FAMILY : IEC
NAME : IEC_TMR
VERSION : 1.0
"IEC_TIMER"
BEGIN
END_DATA_BLOCK

DATA_BLOCK "C11_Heartbeat_On_Timer"   // DB30
{ S7_Optimized_Access := 'TRUE' }
AUTHOR : Simatic
FAMILY : IEC
NAME : IEC_TMR
VERSION : 1.0
"IEC_TIMER"
BEGIN
END_DATA_BLOCK

DATA_BLOCK "C11_Heartbeat_Off_Timer"   // DB31
{ S7_Optimized_Access := 'TRUE' }
AUTHOR : Simatic
FAMILY : IEC
NAME : IEC_TMR
VERSION : 1.0
"IEC_TIMER"
BEGIN
END_DATA_BLOCK

DATA_BLOCK "C12_Heartbeat_On_Timer"   // DB32
{ S7_Optimized_Access := 'TRUE' }
AUTHOR : Simatic
FAMILY : IEC
NAME : IEC_TMR
VERSION : 1.0
"IEC_TIMER"
BEGIN
END_DATA_BLOCK

DATA_BLOCK "C12_Heartbeat_Off_Timer"   // DB33
{ S7_Optimized_Access := 'TRUE' }
AUTHOR : Simatic
FAMILY : IEC
NAME : IEC_TMR
VERSION : 1.0
"IEC_TIMER"
BEGIN
END_DATA_BLOCK

DATA_BLOCK "C13_Heartbeat_On_Timer"   // DB34
{ S7_Optimized_Access := 'TRUE' }
AUTHOR : Simatic
FAMILY : IEC
NAME : IEC_TMR
VERSION : 1.0
"IEC_TIMER"
BEGIN
END_DATA_BLOCK

DATA_BLOCK "C13_Heartbeat_Off_Timer"   // DB35
{ S7_Optimized_Access := 'TRUE' }
AUTHOR : Simatic
FAMILY : IEC
NAME : IEC_TMR
VERSION : 1.0
"IEC_TIMER"
BEGIN
END_DATA_BLOCK

DATA_BLOCK "C14_Heartbeat_On_Timer"   // DB36
{ S7_Optimized_Access := 'TRUE' }
AUTHOR : Simatic
FAMILY : IEC
NAME : IEC_TMR
VERSION : 1.0
"IEC_TIMER"
BEGIN
END_DATA_BLOCK

DATA_BLOCK "C14_Heartbeat_Off_Timer"   // DB37
{ S7_Optimized_Access := 'TRUE' }
AUTHOR : Simatic
FAMILY : IEC
NAME : IEC_TMR
VERSION : 1.0
"IEC_TIMER"
BEGIN
END_DATA_BLOCK

DATA_BLOCK "C15_Heartbeat_On_Timer"   // DB38
{ S7_Optimized_Access := 'TRUE' }
AUTHOR : Simatic
FAMILY : IEC
NAME : IEC_TMR
VERSION : 1.0
"IEC_TIMER"
BEGIN
END_DATA_BLOCK

DATA_BLOCK "C15_Heartbeat_Off_Timer"   // DB39
{ S7_Optimized_Access := 'TRUE' }
AUTHOR : Simatic
FAMILY : IEC
NAME : IEC_TMR
VERSION : 1.0
"IEC_TIMER"
BEGIN
END_DATA_BLOCK

DATA_BLOCK "C16_Heartbeat_On_Timer"   // DB40
{ S7_Optimized_Access := 'TRUE' }
AUTHOR : Simatic
FAMILY : IEC
NAME : IEC_TMR
VERSION : 1.0
"IEC_TIMER"
BEGIN
END_DATA_BLOCK

DATA_BLOCK "C16_Heartbeat_Off_Timer"   // DB41
{ S7_Optimized_Access := 'TRUE' }
AUTHOR : Simatic
FAMILY : IEC
NAME : IEC_TMR
VERSION : 1.0
"IEC_TIMER"
BEGIN
END_DATA_BLOCK

DATA_BLOCK "C17_Heartbeat_On_Timer"   // DB42
{ S7_Optimized_Access := 'TRUE' }
AUTHOR : Simatic
FAMILY : IEC
NAME : IEC_TMR
VERSION : 1.0
"IEC_TIMER"
BEGIN
END_DATA_BLOCK

DATA_BLOCK "C17_Heartbeat_Off_Timer"   // DB43
{ S7_Optimized_Access := 'TRUE' }
AUTHOR : Simatic
FAMILY : IEC
NAME : IEC_TMR
VERSION : 1.0
"IEC_TIMER"
BEGIN
END_DATA_BLOCK

DATA_BLOCK "C18_Heartbeat_On_Timer"   // DB44
{ S7_Optimized_Access := 'TRUE' }
AUTHOR : Simatic
FAMILY : IEC
NAME : IEC_TMR
VERSION : 1.0
"IEC_TIMER"
BEGIN
END_DATA_BLOCK

DATA_BLOCK "C18_Heartbeat_Off_Timer"   // DB45
{ S7_Optimized_Access := 'TRUE' }
AUTHOR : Simatic
FAMILY : IEC
NAME : IEC_TMR
VERSION : 1.0
"IEC_TIMER"
BEGIN
END_DATA_BLOCK

DATA_BLOCK "C19_Heartbeat_On_Timer"   // DB46
{ S7_Optimized_Access := 'TRUE' }
AUTHOR : Simatic
FAMILY : IEC
NAME : IEC_TMR
VERSION : 1.0
"IEC_TIMER"
BEGIN
END_DATA_BLOCK

DATA_BLOCK "C19_Heartbeat_Off_Timer"   // DB47
{ S7_Optimized_Access := 'TRUE' }
AUTHOR : Simatic
FAMILY : IEC
NAME : IEC_TMR
VERSION : 1.0
"IEC_TIMER"
BEGIN
END_DATA_BLOCK

DATA_BLOCK "C20_Heartbeat_On_Timer"   // DB48
{ S7_Optimized_Access := 'TRUE' }
AUTHOR : Simatic
FAMILY : IEC
NAME : IEC_TMR
VERSION : 1.0
"IEC_TIMER"
BEGIN
END_DATA_BLOCK

DATA_BLOCK "C20_Heartbeat_Off_Timer"   // DB49
{ S7_Optimized_Access := 'TRUE' }
AUTHOR : Simatic
FAMILY : IEC
NAME : IEC_TMR
VERSION : 1.0
"IEC_TIMER"
BEGIN
END_DATA_BLOCK

DATA_BLOCK "C30_Heartbeat_Off_Timer"   // DB50
{ S7_Optimized_Access := 'TRUE' }
AUTHOR : Simatic
FAMILY : IEC
NAME : IEC_TMR
VERSION : 1.0
"IEC_TIMER"
BEGIN
END_DATA_BLOCK

DATA_BLOCK "C01_Heartbeat_On_Timer"   // DB51
{ S7_Optimized_Access := 'TRUE' }
AUTHOR : Simatic
FAMILY : IEC
NAME : IEC_TMR
VERSION : 1.0
"IEC_TIMER"
BEGIN
END_DATA_BLOCK

DATA_BLOCK "C01_Heartbeat_Off_Timer"   // DB52
{ S7_Optimized_Access := 'TRUE' }
AUTHOR : Simatic
FAMILY : IEC
NAME : IEC_TMR
VERSION : 1.0
"IEC_TIMER"
BEGIN
END_DATA_BLOCK

DATA_BLOCK "C02_Heartbeat_On_Timer"   // DB54
{ S7_Optimized_Access := 'TRUE' }
AUTHOR : Simatic
FAMILY : IEC
NAME : IEC_TMR
VERSION : 1.0
"IEC_TIMER"
BEGIN
END_DATA_BLOCK

DATA_BLOCK "C02_Heartbeat_Off_Timer"   // DB55
{ S7_Optimized_Access := 'TRUE' }
AUTHOR : Simatic
FAMILY : IEC
NAME : IEC_TMR
VERSION : 1.0
"IEC_TIMER"
BEGIN
END_DATA_BLOCK

DATA_BLOCK "C03_Heartbeat_On_Timer"   // DB56
{ S7_Optimized_Access := 'TRUE' }
AUTHOR : Simatic
FAMILY : IEC
NAME : IEC_TMR
VERSION : 1.0
"IEC_TIMER"
BEGIN
END_DATA_BLOCK

DATA_BLOCK "C03_Heartbeat_Off_Timer"   // DB57
{ S7_Optimized_Access := 'TRUE' }
AUTHOR : Simatic
FAMILY : IEC
NAME : IEC_TMR
VERSION : 1.0
"IEC_TIMER"
BEGIN
END_DATA_BLOCK

DATA_BLOCK "C04_Heartbeat_On_Timer"   // DB58
{ S7_Optimized_Access := 'TRUE' }
AUTHOR : Simatic
FAMILY : IEC
NAME : IEC_TMR
VERSION : 1.0
"IEC_TIMER"
BEGIN
END_DATA_BLOCK

DATA_BLOCK "C04_Heartbeat_Off_Timer"   // DB59
{ S7_Optimized_Access := 'TRUE' }
AUTHOR : Simatic
FAMILY : IEC
NAME : IEC_TMR
VERSION : 1.0
"IEC_TIMER"
BEGIN
END_DATA_BLOCK

DATA_BLOCK "C05_Heartbeat_On_Timer"   // DB60
{ S7_Optimized_Access := 'TRUE' }
AUTHOR : Simatic
FAMILY : IEC
NAME : IEC_TMR
VERSION : 1.0
"IEC_TIMER"
BEGIN
END_DATA_BLOCK

DATA_BLOCK "C05_Heartbeat_Off_Timer"   // DB61
{ S7_Optimized_Access := 'TRUE' }
AUTHOR : Simatic
FAMILY : IEC
NAME : IEC_TMR
VERSION : 1.0
"IEC_TIMER"
BEGIN
END_DATA_BLOCK

DATA_BLOCK "C06_Heartbeat_On_Timer"   // DB62
{ S7_Optimized_Access := 'TRUE' }
AUTHOR : Simatic
FAMILY : IEC
NAME : IEC_TMR
VERSION : 1.0
"IEC_TIMER"
BEGIN
END_DATA_BLOCK

DATA_BLOCK "C06_Heartbeat_Off_Timer"   // DB63
{ S7_Optimized_Access := 'TRUE' }
AUTHOR : Simatic
FAMILY : IEC
NAME : IEC_TMR
VERSION : 1.0
"IEC_TIMER"
BEGIN
END_DATA_BLOCK

DATA_BLOCK "C07_Heartbeat_On_Timer"   // DB64
{ S7_Optimized_Access := 'TRUE' }
AUTHOR : Simatic
FAMILY : IEC
NAME : IEC_TMR
VERSION : 1.0
"IEC_TIMER"
BEGIN
END_DATA_BLOCK

DATA_BLOCK "C07_Heartbeat_Off_Timer"   // DB65
{ S7_Optimized_Access := 'TRUE' }
AUTHOR : Simatic
FAMILY : IEC
NAME : IEC_TMR
VERSION : 1.0
"IEC_TIMER"
BEGIN
END_DATA_BLOCK

DATA_BLOCK "C08_Heartbeat_On_Timer"   // DB66
{ S7_Optimized_Access := 'TRUE' }
AUTHOR : Simatic
FAMILY : IEC
NAME : IEC_TMR
VERSION : 1.0
"IEC_TIMER"
BEGIN
END_DATA_BLOCK

DATA_BLOCK "C08_Heartbeat_Off_Timer"   // DB67
{ S7_Optimized_Access := 'TRUE' }
AUTHOR : Simatic
FAMILY : IEC
NAME : IEC_TMR
VERSION : 1.0
"IEC_TIMER"
BEGIN
END_DATA_BLOCK

DATA_BLOCK "C09_Heartbeat_On_Timer"   // DB68
{ S7_Optimized_Access := 'TRUE' }